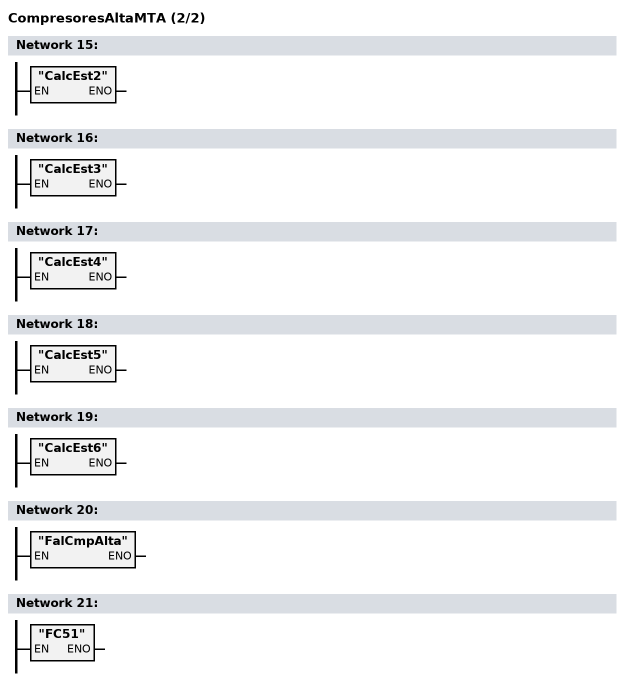
   RUNG wire#powerrail
      "CalcEst2"()
   END_RUNG
   // the same network as SCL:
   "CalcEst2"();
END_REGION

REGION Network 16
   RUNG wire#powerrail
      "CalcEst3"()
   END_RUNG
   // the same network as SCL:
   "CalcEst3"();
END_REGION

REGION Network 17
   RUNG wire#powerrail
      "CalcEst4"()
   END_RUNG
   // the same network as SCL:
   "CalcEst4"();
END_REGION

REGION Network 18
   RUNG wire#powerrail
      "CalcEst5"()
   END_RUNG
   // the same network as SCL:
   "CalcEst5"();
END_REGION

REGION Network 19
   RUNG wire#powerrail
      "CalcEst6"()
   END_RUNG
   // the same network as SCL:
   "CalcEst6"();
END_REGION

REGION Network 20
   RUNG wire#powerrail
      "FalCmpAlta"()
   END_RUNG
   // the same network as SCL:
   "FalCmpAlta"();
END_REGION

REGION Network 21
   RUNG wire#powerrail
      "FC51"()
   END_RUNG
   // the same network as SCL:
   "FC51"();
END_REGION
END_FUNCTION

FUNCTION "ParamCmpALTA-MTA" : Void   // FC30, LAD
{ S7_Optimized_Access := 'FALSE' }
VERSION : 0.1
BEGIN

REGION Network 1
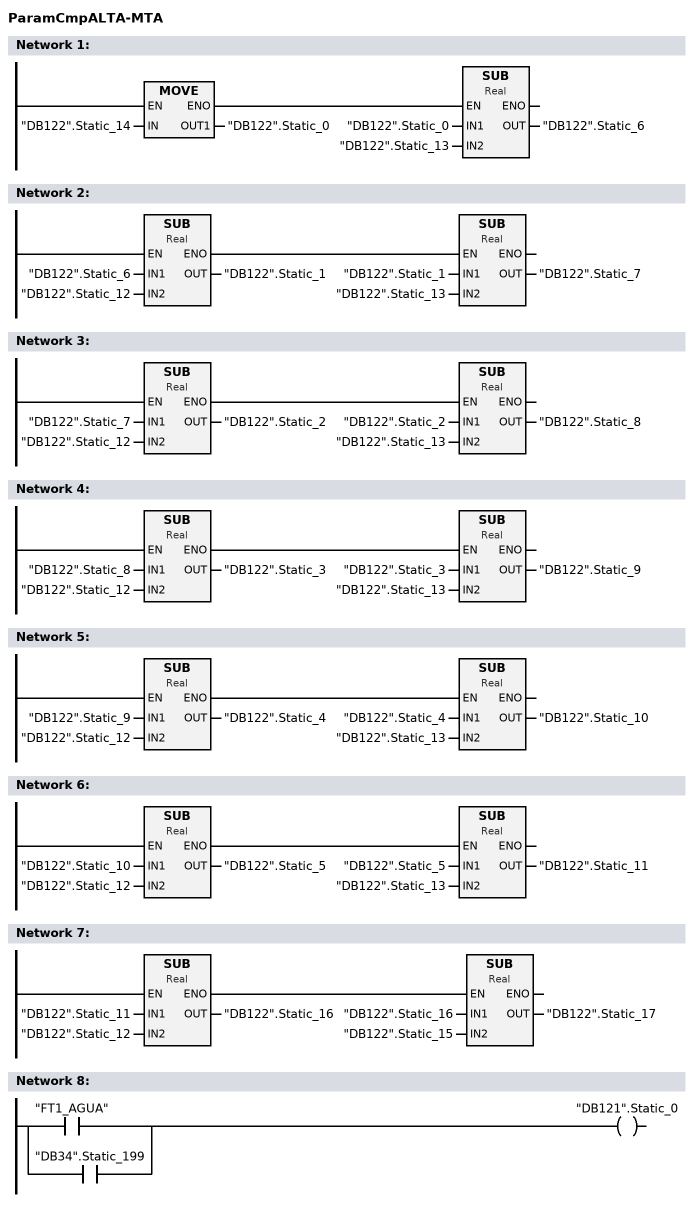
   RUNG wire#powerrail
      { S7_GenerateENO := "TRUE" } Move(in := "DB122".Static_14, out1 => "DB122".Static_0)
      { S7_Templates := "SrcType := Real"; S7_GenerateENO := "TRUE" } Sub(in1 := "DB122".Static_0, in2 := "DB122".Static_13, out => "DB122".Static_6)
   END_RUNG
   // the same network as SCL:
   // ENO of a box is taken as its EN; it also drops when the box reports an error
   "DB122".Static_0 := "DB122".Static_14;
   "DB122".Static_6 := "DB122".Static_0 - "DB122".Static_13;
END_REGION

REGION Network 2
   RUNG wire#powerrail
      { S7_Templates := "SrcType := Real"; S7_GenerateENO := "TRUE" } Sub(in1 := "DB122".Static_6, in2 := "DB122".Static_12, out => "DB122".Static_1)
      { S7_Templates := "SrcType := Real"; S7_GenerateENO := "TRUE" } Sub(in1 := "DB122".Static_1, in2 := "DB122".Static_13, out => "DB122".Static_7)
   END_RUNG
   // the same network as SCL:
   // ENO of a box is taken as its EN; it also drops when the box reports an error
   "DB122".Static_1 := "DB122".Static_6 - "DB122".Static_12;
   "DB122".Static_7 := "DB122".Static_1 - "DB122".Static_13;
END_REGION

REGION Network 3
   RUNG wire#powerrail
      { S7_Templates := "SrcType := Real"; S7_GenerateENO := "TRUE" } Sub(in1 := "DB122".Static_7, in2 := "DB122".Static_12, out => "DB122".Static_2)
      { S7_Templates := "SrcType := Real"; S7_GenerateENO := "TRUE" } Sub(in1 := "DB122".Static_2, in2 := "DB122".Static_13, out => "DB122".Static_8)
   END_RUNG
   // the same network as SCL:
   // ENO of a box is taken as its EN; it also drops when the box reports an error
   "DB122".Static_2 := "DB122".Static_7 - "DB122".Static_12;
   "DB122".Static_8 := "DB122".Static_2 - "DB122".Static_13;
END_REGION

REGION Network 4
   RUNG wire#powerrail
      { S7_Templates := "SrcType := Real"; S7_GenerateENO := "TRUE" } Sub(in1 := "DB122".Static_8, in2 := "DB122".Static_12, out => "DB122".Static_3)
      { S7_Templates := "SrcType := Real"; S7_GenerateENO := "TRUE" } Sub(in1 := "DB122".Static_3, in2 := "DB122".Static_13, out => "DB122".Static_9)
   END_RUNG
   // the same network as SCL:
   // ENO of a box is taken as its EN; it also drops when the box reports an error
   "DB122".Static_3 := "DB122".Static_8 - "DB122".Static_12;
   "DB122".Static_9 := "DB122".Static_3 - "DB122".Static_13;
END_REGION

REGION Network 5
   RUNG wire#powerrail
      { S7_Templates := "SrcType := Real"; S7_GenerateENO := "TRUE" } Sub(in1 := "DB122".Static_9, in2 := "DB122".Static_12, out => "DB122".Static_4)
      { S7_Templates := "SrcType := Real"; S7_GenerateENO := "TRUE" } Sub(in1 := "DB122".Static_4, in2 := "DB122".Static_13, out => "DB122".Static_10)
   END_RUNG
   // the same network as SCL:
   // ENO of a box is taken as its EN; it also drops when the box reports an error
   "DB122".Static_4 := "DB122".Static_9 - "DB122".Static_12;
   "DB122".Static_10 := "DB122".Static_4 - "DB122".Static_13;
END_REGION

REGION Network 6
   RUNG wire#powerrail
      { S7_Templates := "SrcType := Real"; S7_GenerateENO := "TRUE" } Sub(in1 := "DB122".Static_10, in2 := "DB122".Static_12, out => "DB122".Static_5)
      { S7_Templates := "SrcType := Real"; S7_GenerateENO := "TRUE" } Sub(in1 := "DB122".Static_5, in2 := "DB122".Static_13, out => "DB122".Static_11)
   END_RUNG
   // the same network as SCL:
   // ENO of a box is taken as its EN; it also drops when the box reports an error
   "DB122".Static_5 := "DB122".Static_10 - "DB122".Static_12;
   "DB122".Static_11 := "DB122".Static_5 - "DB122".Static_13;
END_REGION

REGION Network 7
   RUNG wire#powerrail
      { S7_Templates := "SrcType := Real"; S7_GenerateENO := "TRUE" } Sub(in1 := "DB122".Static_11, in2 := "DB122".Static_12, out => "DB122".Static_16)
      { S7_Templates := "SrcType := Real"; S7_GenerateENO := "TRUE" } Sub(in1 := "DB122".Static_16, in2 := "DB122".Static_15, out => "DB122".Static_17)
   END_RUNG
   // the same network as SCL:
   // ENO of a box is taken as its EN; it also drops when the box reports an error
   "DB122".Static_16 := "DB122".Static_11 - "DB122".Static_12;
   "DB122".Static_17 := "DB122".Static_16 - "DB122".Static_15;
END_REGION

REGION Network 8
   RUNG wire#powerrail
      Contact( "FT1_AGUA" )
      wire#w1
      Coil( "DB121".Static_0 )
   END_RUNG
   RUNG wire#powerrail
      Contact( "DB34".Static_199 )
   END_RUNG wire#w1
   // the same network as SCL:
   "DB121".Static_0 := "FT1_AGUA" OR "DB34".Static_199;
END_REGION
END_FUNCTION

FUNCTION "TiemposCMPAlta-MTA" : Void   // FC31, LAD
{ S7_Optimized_Access := 'FALSE' }
VERSION : 0.1
   VAR_TEMP   // added for the SCL form of the ladder/FBD networks
      _s5time1 : S5Time;
   END_VAR
BEGIN

REGION Network 1
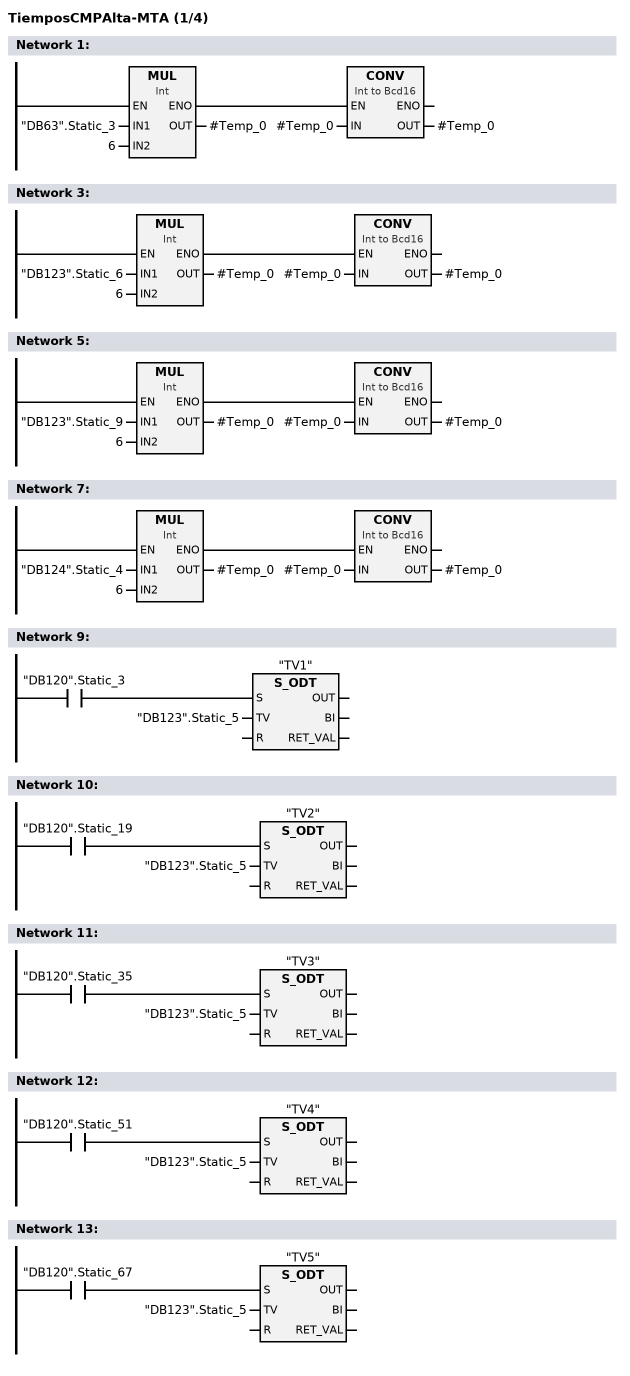
   RUNG wire#powerrail
      { S7_Templates := "SrcType := Int"; S7_GenerateENO := "TRUE" } Mul(in1 := "DB63".Static_3, in2 := 6, out => #Temp_0)
      { S7_Templates := "[SrcType := Int, DestType := Bcd16]"; S7_GenerateENO := "TRUE" } Convert(in := #Temp_0, out => #Temp_0)
   END_RUNG
   // the same network as SCL:
   // ENO of a box is taken as its EN; it also drops when the box reports an error
   #Temp_0 := "DB63".Static_3 * 6;
   #Temp_0 := INT_TO_BCD16(#Temp_0);
END_REGION

REGION Network 2 (STL)
         L     12288;
         L     #Temp_0;
         OW;
         T     "DB63".Static_0;
         NOP   0;
END_REGION

REGION Network 3
   RUNG wire#powerrail
      { S7_Templates := "SrcType := Int"; S7_GenerateENO := "TRUE" } Mul(in1 := "DB123".Static_6, in2 := 6, out => #Temp_0)
      { S7_Templates := "[SrcType := Int, DestType := Bcd16]"; S7_GenerateENO := "TRUE" } Convert(in := #Temp_0, out => #Temp_0)
   END_RUNG
   // the same network as SCL:
   // ENO of a box is taken as its EN; it also drops when the box reports an error
   #Temp_0 := "DB123".Static_6 * 6;
   #Temp_0 := INT_TO_BCD16(#Temp_0);
END_REGION

REGION Network 4 (STL)
         L     12288;
         L     #Temp_0;
         OW;
         T     "DB123".Static_5;
         NOP   0;
END_REGION

REGION Network 5
   RUNG wire#powerrail
      { S7_Templates := "SrcType := Int"; S7_GenerateENO := "TRUE" } Mul(in1 := "DB123".Static_9, in2 := 6, out => #Temp_0)
      { S7_Templates := "[SrcType := Int, DestType := Bcd16]"; S7_GenerateENO := "TRUE" } Convert(in := #Temp_0, out => #Temp_0)
   END_RUNG
   // the same network as SCL:
   // ENO of a box is taken as its EN; it also drops when the box reports an error
   #Temp_0 := "DB123".Static_9 * 6;
   #Temp_0 := INT_TO_BCD16(#Temp_0);
END_REGION

REGION Network 6 (STL)
         L     12288;
         L     #Temp_0;
         OW;
         T     "DB123".Static_8;
         NOP   0;
END_REGION

REGION Network 7
   RUNG wire#powerrail
      { S7_Templates := "SrcType := Int"; S7_GenerateENO := "TRUE" } Mul(in1 := "DB124".Static_4, in2 := 6, out => #Temp_0)
      { S7_Templates := "[SrcType := Int, DestType := Bcd16]"; S7_GenerateENO := "TRUE" } Convert(in := #Temp_0, out => #Temp_0)
   END_RUNG
   // the same network as SCL:
   // ENO of a box is taken as its EN; it also drops when the box reports an error
   #Temp_0 := "DB124".Static_4 * 6;
   #Temp_0 := INT_TO_BCD16(#Temp_0);
END_REGION

REGION Network 8 (STL)
         L     12288;
         L     #Temp_0;
         OW;
         T     "DB124".Static_3;
         NOP   0;
END_REGION

REGION Network 9
   RUNG wire#powerrail
      Contact( "DB120".Static_3 )
      S_ODT(T_NO := "TV1", TV := "DB123".Static_5, R :=, BI =>, RET_VAL =>)
   END_RUNG
   // the same network as SCL:
   #_s5time1 := S_ODT(T_NO := "TV1", TV := "DB123".Static_5, S := "DB120".Static_3);
END_REGION

REGION Network 10
   RUNG wire#powerrail
      Contact( "DB120".Static_19 )
      S_ODT(T_NO := "TV2", TV := "DB123".Static_5, R :=, BI =>, RET_VAL =>)
   END_RUNG
   // the same network as SCL:
   #_s5time1 := S_ODT(T_NO := "TV2", TV := "DB123".Static_5, S := "DB120".Static_19);
END_REGION

REGION Network 11
   RUNG wire#powerrail
      Contact( "DB120".Static_35 )
      S_ODT(T_NO := "TV3", TV := "DB123".Static_5, R :=, BI =>, RET_VAL =>)
   END_RUNG
   // the same network as SCL:
   #_s5time1 := S_ODT(T_NO := "TV3", TV := "DB123".Static_5, S := "DB120".Static_35);
END_REGION

REGION Network 12
   RUNG wire#powerrail
      Contact( "DB120".Static_51 )
      S_ODT(T_NO := "TV4", TV := "DB123".Static_5, R :=, BI =>, RET_VAL =>)
   END_RUNG
   // the same network as SCL:
   #_s5time1 := S_ODT(T_NO := "TV4", TV := "DB123".Static_5, S := "DB120".Static_51);
END_REGION

REGION Network 13
   RUNG wire#powerrail
      Contact( "DB120".Static_67 )
      S_ODT(T_NO := "TV5", TV := "DB123".Static_5, R :=, BI =>, RET_VAL =>)
   END_RUNG
   // the same network as SCL:
   #_s5time1 := S_ODT(T_NO := "TV5", TV := "DB123".Static_5, S := "DB120".Static_67);
END_REGION

REGION Network 14
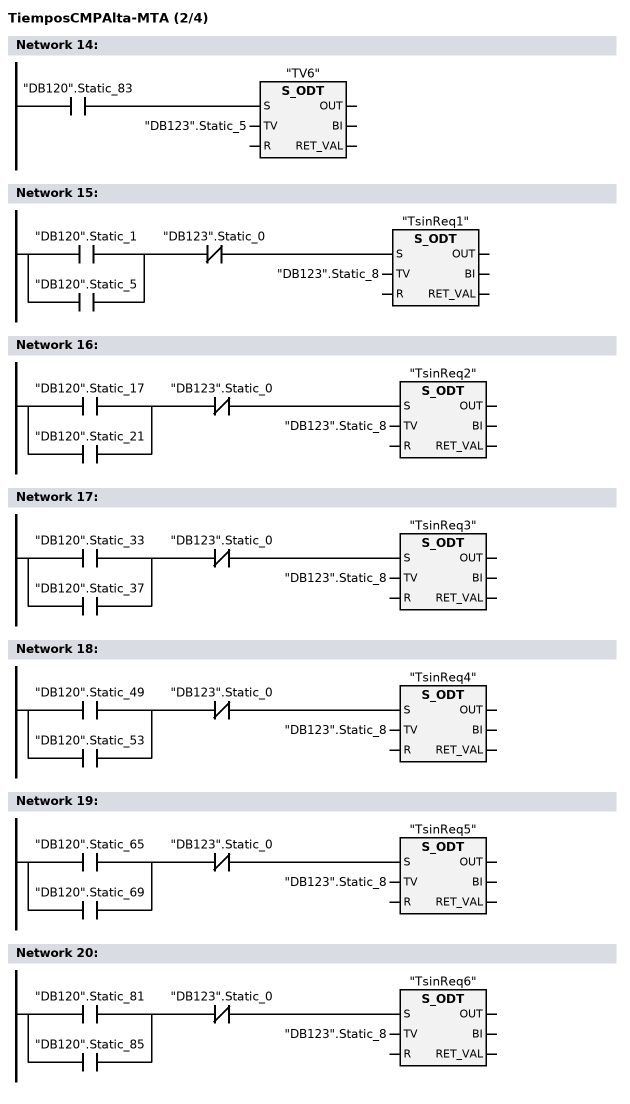
   RUNG wire#powerrail
      Contact( "DB120".Static_83 )
      S_ODT(T_NO := "TV6", TV := "DB123".Static_5, R :=, BI =>, RET_VAL =>)
   END_RUNG
   // the same network as SCL:
   #_s5time1 := S_ODT(T_NO := "TV6", TV := "DB123".Static_5, S := "DB120".Static_83);
END_REGION

REGION Network 15
   RUNG wire#powerrail
      Contact( "DB120".Static_1 )
      wire#w1
      I_Contact( "DB123".Static_0 )
      S_ODT(T_NO := "TsinReq1", TV := "DB123".Static_8, R :=, BI =>, RET_VAL =>)
   END_RUNG
   RUNG wire#powerrail
      Contact( "DB120".Static_5 )
   END_RUNG wire#w1
   // the same network as SCL:
   #_s5time1 := S_ODT(T_NO := "TsinReq1",
                      TV := "DB123".Static_8,
                      S := ("DB120".Static_1 OR "DB120".Static_5) AND NOT "DB123".Static_0);
END_REGION

REGION Network 16
   RUNG wire#powerrail
      Contact( "DB120".Static_17 )
      wire#w1
      I_Contact( "DB123".Static_0 )
      S_ODT(T_NO := "TsinReq2", TV := "DB123".Static_8, R :=, BI =>, RET_VAL =>)
   END_RUNG
   RUNG wire#powerrail
      Contact( "DB120".Static_21 )
   END_RUNG wire#w1
   // the same network as SCL:
   #_s5time1 := S_ODT(T_NO := "TsinReq2",
                      TV := "DB123".Static_8,
                      S := ("DB120".Static_17 OR "DB120".Static_21) AND NOT "DB123".Static_0);
END_REGION

REGION Network 17
   RUNG wire#powerrail
      Contact( "DB120".Static_33 )
      wire#w1
      I_Contact( "DB123".Static_0 )
      S_ODT(T_NO := "TsinReq3", TV := "DB123".Static_8, R :=, BI =>, RET_VAL =>)
   END_RUNG
   RUNG wire#powerrail
      Contact( "DB120".Static_37 )
   END_RUNG wire#w1
   // the same network as SCL:
   #_s5time1 := S_ODT(T_NO := "TsinReq3",
                      TV := "DB123".Static_8,
                      S := ("DB120".Static_33 OR "DB120".Static_37) AND NOT "DB123".Static_0);
END_REGION

REGION Network 18
   RUNG wire#powerrail
      Contact( "DB120".Static_49 )
      wire#w1
      I_Contact( "DB123".Static_0 )
      S_ODT(T_NO := "TsinReq4", TV := "DB123".Static_8, R :=, BI =>, RET_VAL =>)
   END_RUNG
   RUNG wire#powerrail
      Contact( "DB120".Static_53 )
   END_RUNG wire#w1
   // the same network as SCL:
   #_s5time1 := S_ODT(T_NO := "TsinReq4",
                      TV := "DB123".Static_8,
                      S := ("DB120".Static_49 OR "DB120".Static_53) AND NOT "DB123".Static_0);
END_REGION

REGION Network 19
   RUNG wire#powerrail
      Contact( "DB120".Static_65 )
      wire#w1
      I_Contact( "DB123".Static_0 )
      S_ODT(T_NO := "TsinReq5", TV := "DB123".Static_8, R :=, BI =>, RET_VAL =>)
   END_RUNG
   RUNG wire#powerrail
      Contact( "DB120".Static_69 )
   END_RUNG wire#w1
   // the same network as SCL:
   #_s5time1 := S_ODT(T_NO := "TsinReq5",
                      TV := "DB123".Static_8,
                      S := ("DB120".Static_65 OR "DB120".Static_69) AND NOT "DB123".Static_0);
END_REGION

REGION Network 20
   RUNG wire#powerrail
      Contact( "DB120".Static_81 )
      wire#w1
      I_Contact( "DB123".Static_0 )
      S_ODT(T_NO := "TsinReq6", TV := "DB123".Static_8, R :=, BI =>, RET_VAL =>)
   END_RUNG
   RUNG wire#powerrail
      Contact( "DB120".Static_85 )
   END_RUNG wire#w1
   // the same network as SCL:
   #_s5time1 := S_ODT(T_NO := "TsinReq6",
                      TV := "DB123".Static_8,
                      S := ("DB120".Static_81 OR "DB120".Static_85) AND NOT "DB123".Static_0);
END_REGION

REGION Network 21
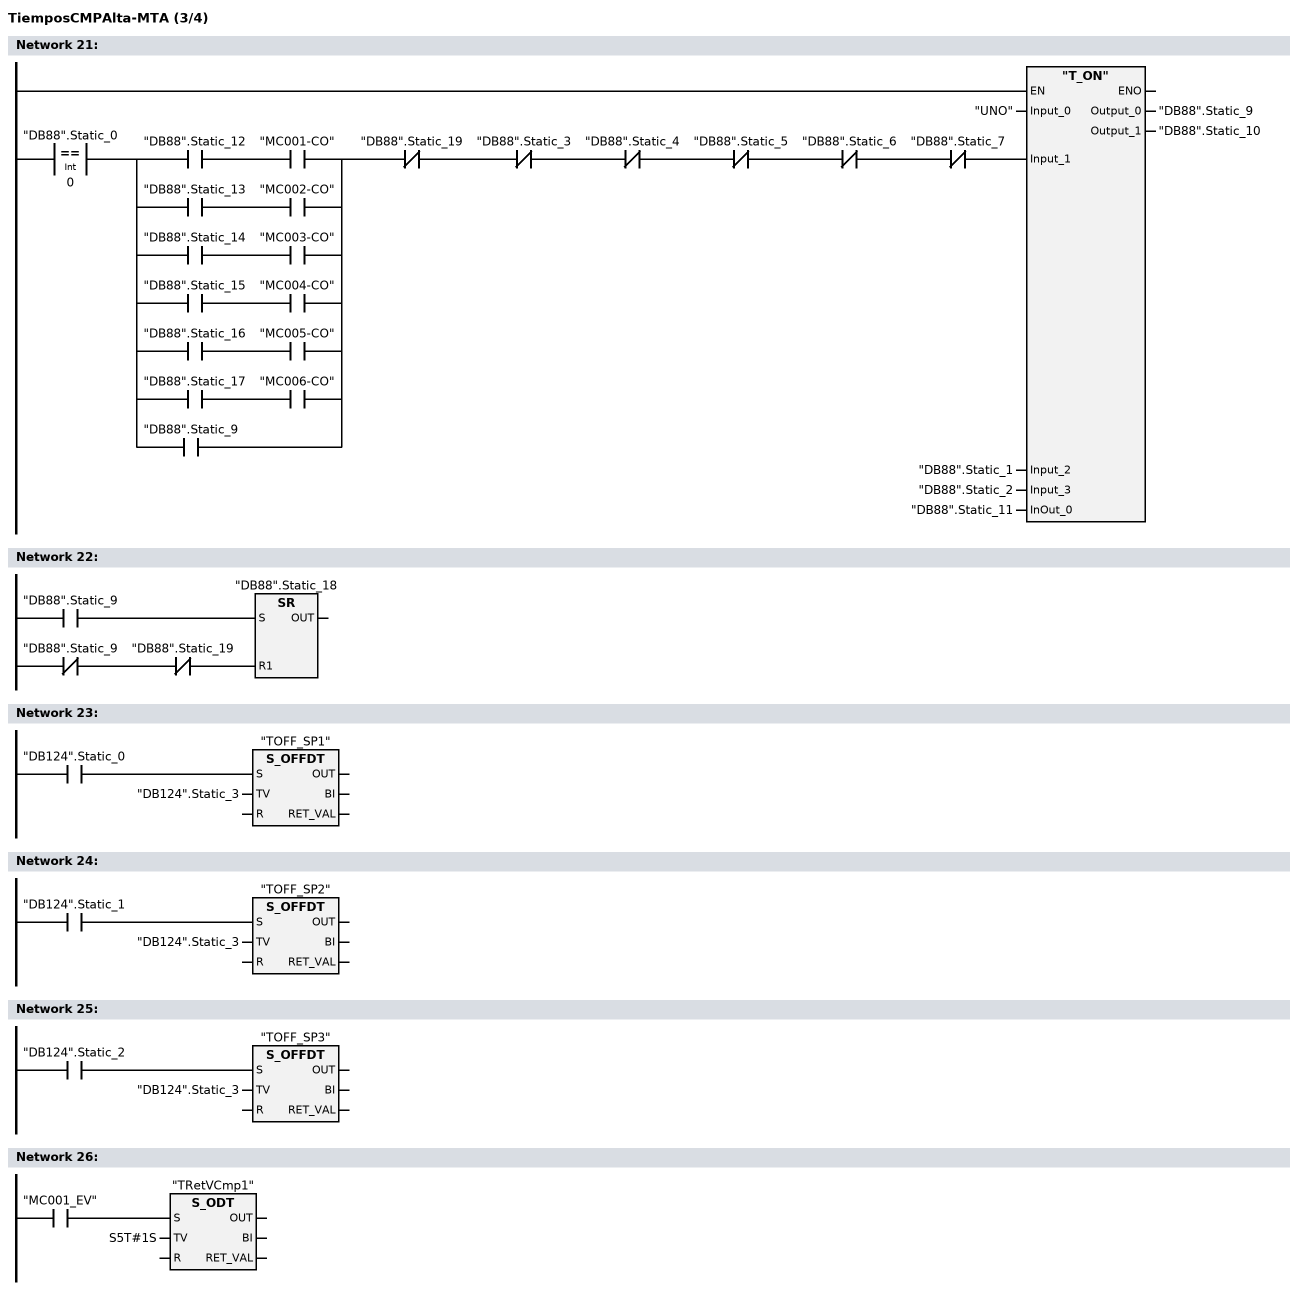
   RUNG wire#powerrail
      "T_ON"(Input_0 := "UNO", Input_2 := "DB88".Static_1, Input_3 := "DB88".Static_2, Output_0 => "DB88".Static_9, Output_1 => "DB88".Static_10, InOut_0 := "DB88".Static_11, Input_1 := wire#w3)
   END_RUNG
   RUNG wire#powerrail
      { S7_Templates := "SrcType := Int" } EQ_Contact(in1 := "DB88".Static_0, in2 := 0)
      wire#w1
      Contact( "DB88".Static_12 )
      Contact( "MC001-CO" )
      wire#w2
      I_Contact( "DB88".Static_19 )
      I_Contact( "DB88".Static_3 )
      I_Contact( "DB88".Static_4 )
      I_Contact( "DB88".Static_5 )
      I_Contact( "DB88".Static_6 )
      I_Contact( "DB88".Static_7 )
   END_RUNG wire#w3
   RUNG wire#w1
      Contact( "DB88".Static_13 )
      Contact( "MC002-CO" )
   END_RUNG wire#w2
   RUNG wire#w1
      Contact( "DB88".Static_14 )
      Contact( "MC003-CO" )
   END_RUNG wire#w2
   RUNG wire#w1
      Contact( "DB88".Static_15 )
      Contact( "MC004-CO" )
   END_RUNG wire#w2
   RUNG wire#w1
      Contact( "DB88".Static_16 )
      Contact( "MC005-CO" )
   END_RUNG wire#w2
   RUNG wire#w1
      Contact( "DB88".Static_17 )
      Contact( "MC006-CO" )
   END_RUNG wire#w2
   RUNG wire#w1
      Contact( "DB88".Static_9 )
   END_RUNG wire#w2
   // the same network as SCL:
   "T_ON"(Input_0 := "UNO",
          Input_1 := ("DB88".Static_0 = 0) AND (("DB88".Static_12 AND "MC001-CO") OR ("DB88".Static_13 AND "MC002-CO") OR ("DB88".Static_14 AND "MC003-CO") OR ("DB88".Static_15 AND "MC004-CO") OR ("DB88".Static_16 AND "MC005-CO") OR ("DB88".Static_17 AND "MC006-CO") OR "DB88".Static_9) AND NOT "DB88".Static_19 AND NOT "DB88".Static_3 AND NOT "DB88".Static_4 AND NOT "DB88".Static_5 AND NOT "DB88".Static_6 AND NOT "DB88".Static_7,
          Input_2 := "DB88".Static_1,
          Input_3 := "DB88".Static_2,
          InOut_0 := "DB88".Static_11,
          Output_0 => "DB88".Static_9,
          Output_1 => "DB88".Static_10);
END_REGION

REGION Network 22
   IF "DB88".Static_9 THEN
       "DB88".Static_18 := TRUE;   // SR flip-flop
   END_IF;
   IF NOT "DB88".Static_9 AND NOT "DB88".Static_19 THEN "DB88".Static_18 := FALSE; END_IF;
END_REGION

REGION Network 23
   RUNG wire#powerrail
      Contact( "DB124".Static_0 )
      S_OFFDT(T_NO := "TOFF_SP1", TV := "DB124".Static_3, R :=, BI =>, RET_VAL =>)
   END_RUNG
   // the same network as SCL:
   #_s5time1 := S_OFFDT(T_NO := "TOFF_SP1", TV := "DB124".Static_3, S := "DB124".Static_0);
END_REGION

REGION Network 24
   RUNG wire#powerrail
      Contact( "DB124".Static_1 )
      S_OFFDT(T_NO := "TOFF_SP2", TV := "DB124".Static_3, R :=, BI =>, RET_VAL =>)
   END_RUNG
   // the same network as SCL:
   #_s5time1 := S_OFFDT(T_NO := "TOFF_SP2", TV := "DB124".Static_3, S := "DB124".Static_1);
END_REGION

REGION Network 25
   RUNG wire#powerrail
      Contact( "DB124".Static_2 )
      S_OFFDT(T_NO := "TOFF_SP3", TV := "DB124".Static_3, R :=, BI =>, RET_VAL =>)
   END_RUNG
   // the same network as SCL:
   #_s5time1 := S_OFFDT(T_NO := "TOFF_SP3", TV := "DB124".Static_3, S := "DB124".Static_2);
END_REGION

REGION Network 26
   RUNG wire#powerrail
      Contact( "MC001_EV" )
      S_ODT(T_NO := "TRetVCmp1", TV := S5T#1S, R :=, BI =>, RET_VAL =>)
   END_RUNG
   // the same network as SCL:
   #_s5time1 := S_ODT(T_NO := "TRetVCmp1", TV := S5T#1S, S := "MC001_EV");
END_REGION

REGION Network 27
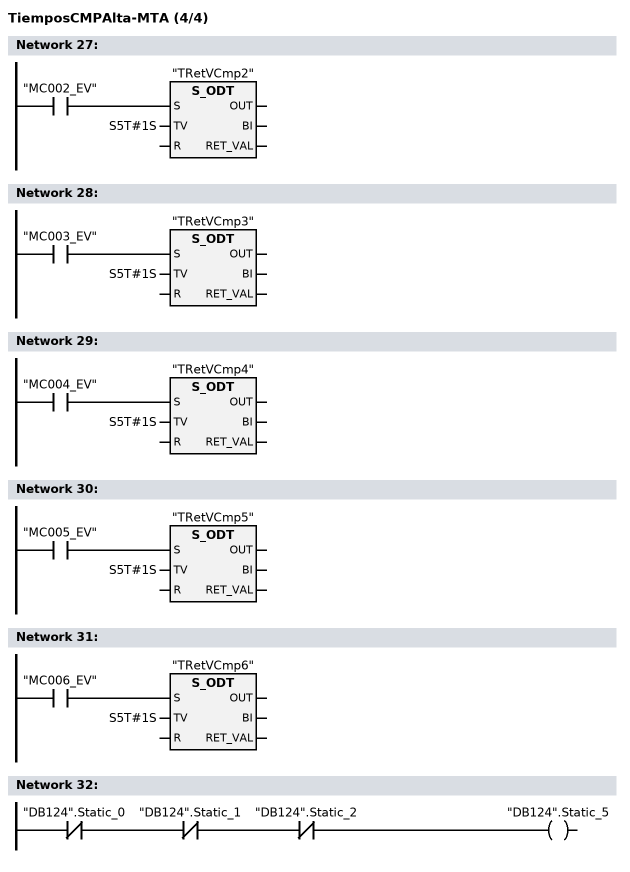
   RUNG wire#powerrail
      Contact( "MC002_EV" )
      S_ODT(T_NO := "TRetVCmp2", TV := S5T#1S, R :=, BI =>, RET_VAL =>)
   END_RUNG
   // the same network as SCL:
   #_s5time1 := S_ODT(T_NO := "TRetVCmp2", TV := S5T#1S, S := "MC002_EV");
END_REGION

REGION Network 28
   RUNG wire#powerrail
      Contact( "MC003_EV" )
      S_ODT(T_NO := "TRetVCmp3", TV := S5T#1S, R :=, BI =>, RET_VAL =>)
   END_RUNG
   // the same network as SCL:
   #_s5time1 := S_ODT(T_NO := "TRetVCmp3", TV := S5T#1S, S := "MC003_EV");
END_REGION

REGION Network 29
   RUNG wire#powerrail
      Contact( "MC004_EV" )
      S_ODT(T_NO := "TRetVCmp4", TV := S5T#1S, R :=, BI =>, RET_VAL =>)
   END_RUNG
   // the same network as SCL:
   #_s5time1 := S_ODT(T_NO := "TRetVCmp4", TV := S5T#1S, S := "MC004_EV");
END_REGION

REGION Network 30
   RUNG wire#powerrail
      Contact( "MC005_EV" )
      S_ODT(T_NO := "TRetVCmp5", TV := S5T#1S, R :=, BI =>, RET_VAL =>)
   END_RUNG
   // the same network as SCL:
   #_s5time1 := S_ODT(T_NO := "TRetVCmp5", TV := S5T#1S, S := "MC005_EV");
END_REGION

REGION Network 31
   RUNG wire#powerrail
      Contact( "MC006_EV" )
      S_ODT(T_NO := "TRetVCmp6", TV := S5T#1S, R :=, BI =>, RET_VAL =>)
   END_RUNG
   // the same network as SCL:
   #_s5time1 := S_ODT(T_NO := "TRetVCmp6", TV := S5T#1S, S := "MC006_EV");
END_REGION

REGION Network 32
   RUNG wire#powerrail
      I_Contact( "DB124".Static_0 )
      I_Contact( "DB124".Static_1 )
      I_Contact( "DB124".Static_2 )
      Coil( "DB124".Static_5 )
   END_RUNG
   // the same network as SCL:
   "DB124".Static_5 := NOT "DB124".Static_0 AND NOT "DB124".Static_1 AND NOT "DB124".Static_2;
END_REGION
END_FUNCTION

FUNCTION "T_ON" : Void   // FC32, LAD
{ S7_Optimized_Access := 'FALSE' }
VERSION : 0.1
   VAR_TEMP   // added for the SCL form of the ladder/FBD networks
      _w1 : Bool;
   END_VAR
BEGIN

REGION Network 1
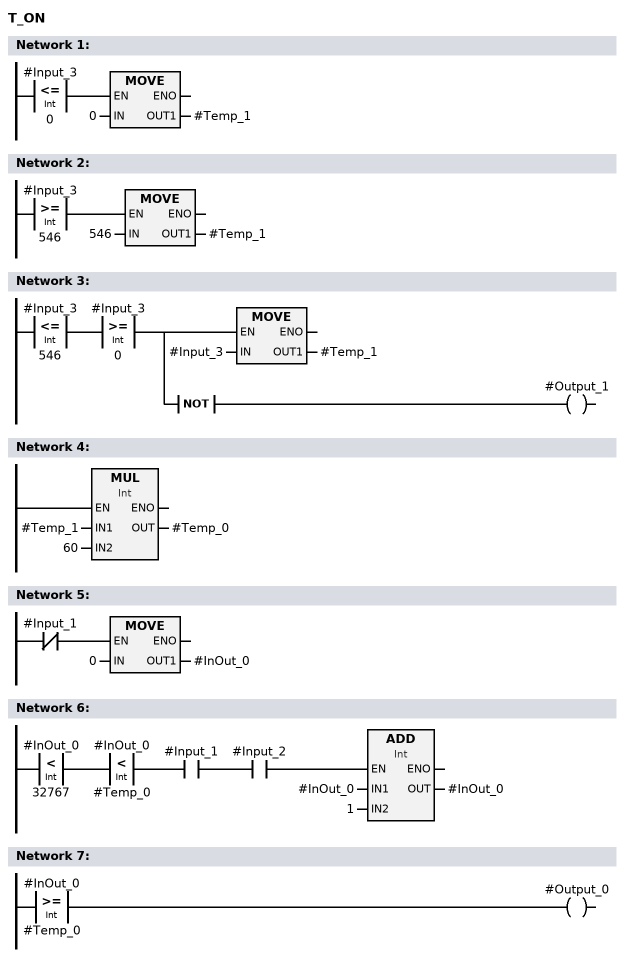
   RUNG wire#powerrail
      { S7_Templates := "SrcType := Int" } LE_Contact(in1 := #Input_3, in2 := 0)
      { S7_GenerateENO := "TRUE" } Move(in := 0, out1 => #Temp_1)
   END_RUNG
   // the same network as SCL:
   IF #Input_3 <= 0 THEN #Temp_1 := 0; END_IF;
END_REGION

REGION Network 2
   RUNG wire#powerrail
      { S7_Templates := "SrcType := Int" } GE_Contact(in1 := #Input_3, in2 := 546)
      { S7_GenerateENO := "TRUE" } Move(in := 546, out1 => #Temp_1)
   END_RUNG
   // the same network as SCL:
   IF #Input_3 >= 546 THEN #Temp_1 := 546; END_IF;
END_REGION

REGION Network 3
   RUNG wire#powerrail
      { S7_Templates := "SrcType := Int" } LE_Contact(in1 := #Input_3, in2 := 546)
      { S7_Templates := "SrcType := Int" } GE_Contact(in1 := #Input_3, in2 := 0)
      wire#w1
      { S7_GenerateENO := "TRUE" } Move(in := #Input_3, out1 => #Temp_1)
   END_RUNG
   RUNG wire#w1
      Not()
      Coil( #Output_1 )
   END_RUNG
   // the same network as SCL:
   #_w1 := (#Input_3 <= 546) AND (#Input_3 >= 0);
   IF #_w1 THEN #Temp_1 := #Input_3; END_IF;
   #Output_1 := NOT #_w1;
END_REGION

REGION Network 4
   RUNG wire#powerrail
      { S7_Templates := "SrcType := Int"; S7_GenerateENO := "TRUE" } Mul(in1 := #Temp_1, in2 := 60, out => #Temp_0)
   END_RUNG
   // the same network as SCL:
   #Temp_0 := #Temp_1 * 60;
END_REGION

REGION Network 5
   RUNG wire#powerrail
      I_Contact( #Input_1 )
      { S7_GenerateENO := "TRUE" } Move(in := 0, out1 => #InOut_0)
   END_RUNG
   // the same network as SCL:
   IF NOT #Input_1 THEN #InOut_0 := 0; END_IF;
END_REGION

REGION Network 6
   RUNG wire#powerrail
      { S7_Templates := "SrcType := Int" } LT_Contact(in1 := #InOut_0, in2 := 32767)
      { S7_Templates := "SrcType := Int" } LT_Contact(in1 := #InOut_0, in2 := #Temp_0)
      Contact( #Input_1 )
      Contact( #Input_2 )
      { S7_Templates := "SrcType := Int"; S7_GenerateENO := "TRUE" } Add(in1 := #InOut_0, in2 := 1, out => #InOut_0)
   END_RUNG
   // the same network as SCL:
   IF (#InOut_0 < 32767) AND (#InOut_0 < #Temp_0) AND #Input_1 AND #Input_2 THEN
       #InOut_0 := #InOut_0 + 1;
   END_IF;
END_REGION

REGION Network 7
   RUNG wire#powerrail
      { S7_Templates := "SrcType := Int" } GE_Contact(in1 := #InOut_0, in2 := #Temp_0)
      Coil( #Output_0 )
   END_RUNG
   // the same network as SCL:
   #Output_0 := #InOut_0 >= #Temp_0;
END_REGION
END_FUNCTION

FUNCTION "PrioridadesCmpAlta" : Void   // FC33, LAD
{ S7_Optimized_Access := 'FALSE' }
VERSION : 0.1
   VAR_TEMP   // added for the SCL form of the ladder/FBD networks
      _w1 : Bool;
   END_VAR
BEGIN

REGION Network 1